// TIA Portal project "E95238_MCC1200_Sisecam_India" (V17)

(* hardware
DEVICE "S71500/ET200MP station_1"  S7-1500 station
   slot 0: "Rail_0"  Rack  6ES7 590-1***0-0AA0
   slot 1: "R150AP1"  CPU 1515-2 PN  6ES7 515-2AM02-0AB0  V2.8
      slot 3: "CPU display_1"  6ES7591-1BA00-0AA0
      slot 32768: "PROFINET_MCC1200"  X1
         slot 32769: "Port_1"  X1 P1
         slot 32770: "Port_2"  X1 P2
      slot 33024: "PCNETWORK_MCC1200"  X2
         slot 33025: "Port_1"  X2 P1
      slot 34817: "Virtual CP interface port_1"  Virtual CP interface port  Virtual CP interface port
   slot 2: "DI 16x24VDC HF_1"  DI 16x24VDC HF  6ES7 521-1BH00-0AB0  V2.2
DEVICE "ET 200SP station_2"  ET 200SP-Station
   slot 0: "Rack_0"  Rack  6ES5 710-8MAx1
   slot 0: "R195AP1"  IM 155-6 PN ST  6ES7 155-6AU01-0BN0  V4.1
   slot 1: "MasterCounter"  TM PosInput 1  6ES7 138-6BA00-0BA0  V1.3
      slot 1: "MasterCounter"  TM PosInput 1
   slot 2: "TM PosInput 1_2"  TM PosInput 1  6ES7 138-6BA00-0BA0  V1.3
      slot 1: "TM PosInput 1_2"  TM PosInput 1
   slot 3: "TM PosInput 1_3"  TM PosInput 1  6ES7 138-6BA00-0BA0  V1.2
      slot 1: "TM PosInput 1_3"  TM PosInput 1
   slot 4: "DI 16x24VDC ST_4"  DI 16x24VDC ST  6ES7 131-6BH01-0BA0  V0.0
      slot 1: "DI 16x24VDC ST_4"  DI 16x24VDC ST
   slot 5: "DI 16x24VDC ST_1"  DI 16x24VDC ST  6ES7 131-6BH01-0BA0  V0.0
      slot 1: "DI 16x24VDC ST_1"  DI 16x24VDC ST
   slot 6: "DI 16x24VDC ST_5"  DI 16x24VDC ST  6ES7 131-6BH01-0BA0  V0.0
      slot 1: "DI 16x24VDC ST_5"  DI 16x24VDC ST
   slot 7: "DQ 16x24VDC/0.5A ST_1"  DQ 16x24VDC/0.5A ST  6ES7 132-6BH01-0BA0  V0.0
      slot 1: "DQ 16x24VDC/0.5A ST_1"  DQ 16x24VDC/0.5A ST
   slot 8: "DQ 16x24VDC/0.5A ST_2"  DQ 16x24VDC/0.5A ST  6ES7 132-6BH01-0BA0  V0.0
      slot 1: "DQ 16x24VDC/0.5A ST_2"  DQ 16x24VDC/0.5A ST
   slot 9: "Server module_1"  Server module  6ES7 193-6PA00-0AA0  V1.1
      slot 1: "Server module_1"  Server module
   slot 127: "BA 2xRJ45"  BA 2xRJ45  6ES7 193-6AR00-0AA0  V0.0
      slot 1: "Port_1"  X1 P1 R  6ES7 193-6AR00-0AA0  V0.0
      slot 2: "Port_2"  X1 P2 R  6ES7 193-6AR00-0AA0  V0.0
DEVICE "ET 200SP station_1"  ET 200SP-Station
   slot 0: "Telaio di montaggio_0"  Rack  6ES5 710-8MAx1
   slot 1: "2B160AP"  CPU 1512SP-1 PN  6ES7 512-1DK01-0AB0  V2.9
      slot 32768: "PROFINET_YC2"  X1
   slot 2: "TM PosInput 1_1"  TM PosInput 1  6ES7 138-6BA00-0BA0  V1.2
      slot 1: "TM PosInput 1_1"  TM PosInput 1
   slot 3: "DI 16x24VDC ST_1"  DI 16x24VDC ST  6ES7 131-6BH01-0BA0  V0.0
      slot 1: "DI 16x24VDC ST_1"  DI 16x24VDC ST
   slot 4: "DI 8x24VDC ST_1"  DI 8x24VDC ST  6ES7 131-6BF01-0BA0  V0.0
      slot 1: "DI 8x24VDC ST_1"  DI 8x24VDC ST
   slot 5: "DQ 8x24VDC/0.5A ST_1"  DQ 8x24VDC/0.5A ST  6ES7 132-6BF01-0BA0  V0.0
      slot 1: "DQ 8x24VDC/0.5A ST_1"  DQ 8x24VDC/0.5A ST
   slot 6: "DQ 8x24VDC/0.5A ST_2"  DQ 8x24VDC/0.5A ST  6ES7 132-6BF01-0BA0  V0.0
      slot 1: "DQ 8x24VDC/0.5A ST_1"  DQ 8x24VDC/0.5A ST
   slot 7: "AQ 4xU/I ST_1"  AQ 4xU/I ST  6ES7 135-6HD00-0BA1  V1.1
      slot 1: "AQ 4xU/I ST_1"  AQ 4xU/I ST
   slot 8: "AQ 4xU/I ST_2"  AQ 4xU/I ST  6ES7 135-6HD00-0BA1  V1.1
      slot 1: "AQ 4xU/I ST_2"  AQ 4xU/I ST
   slot 9: "Modulo server_1"  Server module  6ES7 193-6PA00-0AA0  V1.1
      slot 1: "Modulo server_1"  Server module
   slot 127: "BA 2xRJ45"  BA 2xRJ45  6ES7 193-6AR00-0AA0  V0.0
      slot 32769: "Port_1"  6ES7 193-6AR00-0AA0
      slot 32770: "Port_2"  6ES7 193-6AR00-0AA0
DEVICE "GSD device_1"  GSD.Device.PN
   slot 0: "Rack"  Rack  V1.0
   slot 0: "Y2B412AP1"  55130 IMPACT67 DIO16 IRT  55130  1.02.00
      slot 0: "55130 IMPACT67 DIO16 IRT_1"  55130 IMPACT67 DIO16 IRT
      slot 1: "55130 IMPACT67 DIO16 IRT"  55130 IMPACT67 DIO16 IRT
         slot 1: "Port 1"  Port 1
         slot 2: "Port 2"  Port 2
      slot 1: "Device_1"  Device
         slot 0: "Parameter/Diagnostic"  Parameter/Diagnostic
         slot 1: "Digital IO"  Digital IO
DEVICE "GSD device_3"  GSD.Device.PN
   slot 0: "Rack"  Rack  V1.0
   slot 0: "Y2B411AP1"  55130 IMPACT67 DIO16 IRT  55130  1.02.00
      slot 0: "55130 IMPACT67 DIO16 IRT_1"  55130 IMPACT67 DIO16 IRT
      slot 1: "55130 IMPACT67 DIO16 IRT"  55130 IMPACT67 DIO16 IRT
         slot 1: "Port 1"  Port 1
         slot 2: "Port 2"  Port 2
      slot 1: "Device_1"  Device
         slot 0: "Parameter/Diagnostic"  Parameter/Diagnostic
         slot 1: "Digital IO"  Digital IO
DEVICE "GSD device_4"  GSD.Device.PN
   slot 0: "Rack"  Rack  V1.0
   slot 0: "Y2B413AP1"  55130 IMPACT67 DIO16 IRT  55130  1.02.00
      slot 0: "55130 IMPACT67 DIO16 IRT_1"  55130 IMPACT67 DIO16 IRT
      slot 1: "55130 IMPACT67 DIO16 IRT"  55130 IMPACT67 DIO16 IRT
         slot 1: "Port 1"  Port 1
         slot 2: "Port 2"  Port 2
      slot 1: "Device_1"  Device
         slot 0: "Parameter/Diagnostic"  Parameter/Diagnostic
         slot 1: "Digital IO"  Digital IO
DEVICE "GSD device_5"  GSD.Device.PN
   slot 0: "Rack"  Rack  V1.0
   slot 0: "Y2B414AP1"  55130 IMPACT67 DIO16 IRT  55130  1.02.00
      slot 0: "55130 IMPACT67 DIO16 IRT_1"  55130 IMPACT67 DIO16 IRT
      slot 1: "55130 IMPACT67 DIO16 IRT"  55130 IMPACT67 DIO16 IRT
         slot 1: "Port 1"  Port 1
         slot 2: "Port 2"  Port 2
      slot 1: "Device_1"  Device
         slot 0: "Parameter/Diagnostic"  Parameter/Diagnostic
         slot 1: "Digital IO"  Digital IO
DEVICE "GSD device_7"  GSD.Device.PN
   slot 0: "Rack"  Rack  V1.0
   slot 0: "Y2B415AP1"  55130 IMPACT67 DIO16 IRT  55130  1.02.00
      slot 0: "55130 IMPACT67 DIO16 IRT_1"  55130 IMPACT67 DIO16 IRT
      slot 1: "55130 IMPACT67 DIO16 IRT"  55130 IMPACT67 DIO16 IRT
         slot 1: "Port 1"  Port 1
         slot 2: "Port 2"  Port 2
      slot 1: "Device_1"  Device
         slot 0: "Parameter/Diagnostic"  Parameter/Diagnostic
         slot 1: "Digital IO"  Digital IO
DEVICE "ET 200SP station_3"  ET 200SP-Station
   slot 0: "Telaio di montaggio_0"  Rack  6ES5 710-8MAx1
   slot 1: "1B160AP"  CPU 1512SP-1 PN  6ES7 512-1DK01-0AB0  V2.9
      slot 32768: "PROFINET_YC1"  X1
   slot 2: "TM PosInput 1_1"  TM PosInput 1  6ES7 138-6BA00-0BA0  V1.2
      slot 1: "TM PosInput 1_1"  TM PosInput 1
   slot 3: "DI 16x24VDC ST_1"  DI 16x24VDC ST  6ES7 131-6BH01-0BA0  V0.0
      slot 1: "DI 16x24VDC ST_1"  DI 16x24VDC ST
   slot 4: "DI 8x24VDC ST_1"  DI 8x24VDC ST  6ES7 131-6BF01-0BA0  V0.0
      slot 1: "DI 8x24VDC ST_1"  DI 8x24VDC ST
   slot 5: "DI 16x24VDC ST_2"  DI 16x24VDC ST  6ES7 131-6BH01-0BA0  V0.0
      slot 1: "DI 16x24VDC ST_2"  DI 16x24VDC ST
   slot 6: "DQ 8x24VDC/0.5A ST_1"  DQ 8x24VDC/0.5A ST  6ES7 132-6BF01-0BA0  V0.0
      slot 1: "DQ 8x24VDC/0.5A ST_1"  DQ 8x24VDC/0.5A ST
   slot 7: "DQ 16x24VDC/0.5A ST_1"  DQ 16x24VDC/0.5A ST  6ES7 132-6BH01-0BA0  V0.0
      slot 1: "DQ 16x24VDC/0.5A ST_1"  DQ 16x24VDC/0.5A ST
   slot 8: "AQ 4xU/I ST_1"  AQ 4xU/I ST  6ES7 135-6HD00-0BA1  V1.1
      slot 1: "AQ 4xU/I ST_1"  AQ 4xU/I ST
   slot 9: "AQ 4xU/I ST_2"  AQ 4xU/I ST  6ES7 135-6HD00-0BA1  V1.1
      slot 1: "AQ 4xU/I ST_2"  AQ 4xU/I ST
   slot 10: "Modulo server_1"  Server module  6ES7 193-6PA00-0AA0  V1.1
      slot 1: "Modulo server_1"  Server module
   slot 127: "BA 2xRJ45"  BA 2xRJ45  6ES7 193-6AR00-0AA0  V0.0
      slot 32769: "Port_1"  6ES7 193-6AR00-0AA0
      slot 32770: "Port_2"  6ES7 193-6AR00-0AA0
DEVICE "GSD device_9"  GSD.Device.PN
   slot 0: "Rack"  Rack  V1.0
   slot 0: "Y1B415AP1"  55130 IMPACT67 DIO16 IRT  55130  1.02.00
      slot 0: "55130 IMPACT67 DIO16 IRT_1"  55130 IMPACT67 DIO16 IRT
      slot 1: "55130 IMPACT67 DIO16 IRT"  55130 IMPACT67 DIO16 IRT
         slot 1: "Port 1"  Port 1
         slot 2: "Port 2"  Port 2
      slot 1: "Device_1"  Device
         slot 0: "Parameter/Diagnostic"  Parameter/Diagnostic
         slot 1: "Digital IO"  Digital IO
DEVICE "GSD device_10"  GSD.Device.PN
   slot 0: "Rack"  Rack  V1.0
   slot 0: "Y1B414AP1"  55130 IMPACT67 DIO16 IRT  55130  1.02.00
      slot 0: "55130 IMPACT67 DIO16 IRT_1"  55130 IMPACT67 DIO16 IRT
      slot 1: "55130 IMPACT67 DIO16 IRT"  55130 IMPACT67 DIO16 IRT
         slot 1: "Port 1"  Port 1
         slot 2: "Port 2"  Port 2
      slot 1: "Device_1"  Device
         slot 0: "Parameter/Diagnostic"  Parameter/Diagnostic
         slot 1: "Digital IO"  Digital IO
DEVICE "GSD device_11"  GSD.Device.PN
   slot 0: "Rack"  Rack  V1.0
   slot 0: "Y1B413AP1"  55130 IMPACT67 DIO16 IRT  55130  1.02.00
      slot 0: "55130 IMPACT67 DIO16 IRT_1"  55130 IMPACT67 DIO16 IRT
      slot 1: "55130 IMPACT67 DIO16 IRT"  55130 IMPACT67 DIO16 IRT
         slot 1: "Port 1"  Port 1
         slot 2: "Port 2"  Port 2
      slot 1: "Device_1"  Device
         slot 0: "Parameter/Diagnostic"  Parameter/Diagnostic
         slot 1: "Digital IO"  Digital IO
DEVICE "GSD device_13"  GSD.Device.PN
   slot 0: "Rack"  Rack  V1.0
   slot 0: "Y1B412AP1"  55130 IMPACT67 DIO16 IRT  55130  1.02.00
      slot 0: "55130 IMPACT67 DIO16 IRT_1"  55130 IMPACT67 DIO16 IRT
      slot 1: "55130 IMPACT67 DIO16 IRT"  55130 IMPACT67 DIO16 IRT
         slot 1: "Port 1"  Port 1
         slot 2: "Port 2"  Port 2
      slot 1: "Device_1"  Device
         slot 0: "Parameter/Diagnostic"  Parameter/Diagnostic
         slot 1: "Digital IO"  Digital IO
DEVICE "GSD device_14"  GSD.Device.PN
   slot 0: "Rack"  Rack  V1.0
   slot 0: "Y1B411AP1"  55130 IMPACT67 DIO16 IRT  55130  1.02.00
      slot 0: "55130 IMPACT67 DIO16 IRT_1"  55130 IMPACT67 DIO16 IRT
      slot 1: "55130 IMPACT67 DIO16 IRT"  55130 IMPACT67 DIO16 IRT
         slot 1: "Port 1"  Port 1
         slot 2: "Port 2"  Port 2
      slot 1: "Device_1"  Device
         slot 0: "Parameter/Diagnostic"  Parameter/Diagnostic
         slot 1: "Digital IO"  Digital IO
DEVICE "GSD device_15"  GSD.Device.PN
   slot 0: "Rack"  Rack  V1.0
   slot 0: "Y1B416AP1"  55130 IMPACT67 DIO16 IRT  55130  1.02.00
      slot 0: "55130 IMPACT67 DIO16 IRT_1"  55130 IMPACT67 DIO16 IRT
      slot 1: "55130 IMPACT67 DIO16 IRT"  55130 IMPACT67 DIO16 IRT
         slot 1: "Port 1"  Port 1
         slot 2: "Port 2"  Port 2
      slot 1: "Device_1"  Device
         slot 0: "Parameter/Diagnostic"  Parameter/Diagnostic
         slot 1: "Digital IO"  Digital IO
DEVICE "GSD device_2"  GSD.Device.PN
   slot 0: "Rack"  Rack  V1.0
   slot 0: "Y1B417AP1"  55130 IMPACT67 DIO16 IRT  55130  1.02.00
      slot 0: "55130 IMPACT67 DIO16 IRT_1"  55130 IMPACT67 DIO16 IRT
      slot 1: "55130 IMPACT67 DIO16 IRT"  55130 IMPACT67 DIO16 IRT
         slot 1: "Port 1"  Port 1
         slot 2: "Port 2"  Port 2
      slot 1: "Device_1"  Device
         slot 0: "Parameter/Diagnostic"  Parameter/Diagnostic
         slot 1: "Digital IO"  Digital IO
DEVICE "GSD device_6"  GSD.Device.PN
   slot 0: "Rack"  Rack  V1.0
   slot 0: "Y1B418AP1"  55130 IMPACT67 DIO16 IRT  55130  1.02.00
      slot 0: "55130 IMPACT67 DIO16 IRT_1"  55130 IMPACT67 DIO16 IRT
      slot 1: "55130 IMPACT67 DIO16 IRT"  55130 IMPACT67 DIO16 IRT
         slot 1: "Port 1"  Port 1
         slot 2: "Port 2"  Port 2
      slot 1: "Device_1"  Device
         slot 0: "Parameter/Diagnostic"  Parameter/Diagnostic
         slot 1: "Digital IO"  Digital IO
DEVICE "GSD device_8"  GSD.Device.PN
   slot 0: "Rack"  Rack  V1.0
   slot 0: "Y2B418AP1"  55130 IMPACT67 DIO16 IRT  55130  1.02.00
      slot 0: "55130 IMPACT67 DIO16 IRT_1"  55130 IMPACT67 DIO16 IRT
      slot 1: "55130 IMPACT67 DIO16 IRT"  55130 IMPACT67 DIO16 IRT
         slot 1: "Port 1"  Port 1
         slot 2: "Port 2"  Port 2
      slot 1: "Device_1"  Device
         slot 0: "Parameter/Diagnostic"  Parameter/Diagnostic
         slot 1: "Digital IO"  Digital IO
DEVICE "GSD device_12"  GSD.Device.PN
   slot 0: "Rack"  Rack  V1.0
   slot 0: "Y2B417AP1"  55130 IMPACT67 DIO16 IRT  55130  1.02.00
      slot 0: "55130 IMPACT67 DIO16 IRT_1"  55130 IMPACT67 DIO16 IRT
      slot 1: "55130 IMPACT67 DIO16 IRT"  55130 IMPACT67 DIO16 IRT
         slot 1: "Port 1"  Port 1
         slot 2: "Port 2"  Port 2
      slot 1: "Device_1"  Device
         slot 0: "Parameter/Diagnostic"  Parameter/Diagnostic
         slot 1: "Digital IO"  Digital IO
DEVICE "GSD device_16"  GSD.Device.PN
   slot 0: "Rack"  Rack  V1.0
   slot 0: "Y2B416AP1"  55130 IMPACT67 DIO16 IRT  55130  1.02.00
      slot 0: "55130 IMPACT67 DIO16 IRT_1"  55130 IMPACT67 DIO16 IRT
      slot 1: "55130 IMPACT67 DIO16 IRT"  55130 IMPACT67 DIO16 IRT
         slot 1: "Port 1"  Port 1
         slot 2: "Port 2"  Port 2
      slot 1: "Device_1"  Device
         slot 0: "Parameter/Diagnostic"  Parameter/Diagnostic
         slot 1: "Digital IO"  Digital IO
DEVICE "GSD device_17"  GSD.Device.PN
   slot 0: "Telaio di montaggio"  Rack  V1.0
   slot 1: "d405ap1"  D405AP1  6ES7 512-1DK01-0AB0  V2.9
      slot 0: "InputCPU0"  InputCPU0
      slot 1: "OutputCPU0"  OutputCPU0
      slot 2: "Interface"  Interface
         slot 1: "Port 1"  Port 1
         slot 2: "Port 2"  Port 2
         slot 3: "Port 3"  Port 3
*)

// ===== PLC "R150AP1"  CPU 1515-2 PN =====

VAR_GLOBAL   // PLC tag table "Default tag table"
   "FirstScan" AT %M0.0 : Bool;
   "AlwaysTRUE" AT %M0.2 : Bool;
   "AlwaysFALSE" AT %M0.3 : Bool;
   "AlwaysOFF_Debug" AT %M10.0 : Bool;
   "o.R195AP1.R251KA1.EncoderCommutation" AT %Q120.0 : Bool;
   "i.R195AP1.R11QF2/3.PowerFailure230VAuxiliary" AT %I120.1 : Bool;
   "i.R195AP1.R18QF3.PowerFailure24V_Commands" AT %I120.6 : Bool;
   "i.R195AP1.R18QF4.PowerFailure24V_Input" AT %I120.7 : Bool;
   "i.R195AP1.R18AP1.Redundacy24VOk" AT %I120.5 : Bool;
   "i.R195AP1.M216B1.GlassPresenceOnEncoder#1M216" AT %I122.0 : Bool;
   "i.R195AP1.M216B2.GlassPresenceOnEncoder#2M216" AT %I122.1 : Bool;
   "i.R195AP1.R427SL1.MinimumLevelOilTank" AT %I122.3 : Bool;
   "i.R195AP1.R427SL2.MaximumLevelOilTank" AT %I122.4 : Bool;
   "i.R195AP1.M212SB4.DefectButtonClass3" AT %I123.3 : Bool;
   "i.R195AP1.M212SB3.QualityB1" AT %I123.2 : Bool;
   "i.R195AP1.M212SB5.DefectButtonClass4" AT %I123.4 : Bool;
   "i.R195AP1.SCANNER.ScannerOn" AT %I124.0 : Bool;
   "i.R195AP1.SCANNER.Scanner(1)" AT %I124.1 : Bool;
   "o.R195AP1.R251KA2.Jog" AT %Q120.1 : Bool;
   "o.R195AP1.R252HL1.SafetiesON" AT %Q121.1 : Bool;
   "o.R195AP1.R252HL2.EnableCPUA" AT %Q121.2 : Bool;
   "o.R195AP1.R252HL2.EnableCPUB" AT %Q121.3 : Bool;
   "o.R195AP1.R252KA1.SCANNER.RiseBreakingBar" AT %Q121.5 : Bool;
   "o.R195AP1.R252KA2.SCANNER.GlassToSQC" AT %Q121.6 : Bool;
   "o.R195AP1.M216YV1.DigitizerRise/descentEncoder1" AT %Q122.0 : Bool;
   "o.R195AP1.M216YV2.DigitizeRise/descentEncoder2" AT %Q122.1 : Bool;
   "o.R195AP1.R429YV1.StartFillingPumpCuttingTank" AT %Q122.5 : Bool;
   "o.R195AP1.M221YV2.UpperHolderControl" AT %Q122.7 : Bool;
   "o.R195AP1.M221YV1.BreakoutBarControl" AT %Q122.6 : Bool;
   "o.R195AP1.M221HL1.CutTrasversalBridge1" AT %Q123.1 : Bool;
   "o.R195AP1.M221HL2.CutTrasversalBridge2" AT %Q123.2 : Bool;
   "i.R195AP1.R125KA1CPU_A_Enabled" AT %I121.3 : Bool;
   "i.R195AP1.R125SA1SelectionOnCPU_B" AT %I121.4 : Bool;
   "i.R150AP1.Recognition CPU A" AT %I20.2 : Bool;
   "cigliutti" AT %M100.1 : Bool;
   "i.R195AP1.R18QF7.PowerSupply24VLogic" AT %I121.1 : Bool;
   "i.R195AP1.R427SSP1.CompressedAirPresenceCuttingBridge" AT %I122.5 : Bool;
   "i.R195AP1.R18QF8.PowerSupply24VLogic" AT %I121.2 : Bool;
   "i.R195AP1.M212SB1.DefectButtonClass3" AT %I123.0 : Bool;
   "i.R195AP1.M212SB2.DefectButtonClass4" AT %I123.1 : Bool;
   "o.R195AP1.A255KA6.Anomaly" AT %Q4.5 : Bool;
   "o.R195AP1.A257KA4.AllowM225" AT %Q6.3 : Bool;
   "o.R195AP1.A257KA5.AllowM225(1)" AT %Q6.4 : Bool;
   "o.R195AP1.A252KA3.SCANNER.NoGlassBreak" AT %Q121.7 : Bool;
   "o.R195AP1.M212SB3.M212SB6.GlassRequestQlt" AT %Q123.0 : Bool;
   "o.R195AP1.FanRotationM250" AT %Q2.0 : Bool;
   "i.MCC1256B1_IDevice" AT %I2500.0 : "UDT_YCut_IdeviceFromBridge";
   "i_HSCInput_Count1" AT %I30.0 : "LPD_typeCountFeedbackCh";
   "i_HSCInput_Count2" AT %I160.0 : "LPD_typeCountFeedbackCh";
   "i_HSCInput_Count3" AT %I180.0 : "LPD_typeCountFeedbackCh";
   "i.MCC1256B2_IDevice" AT %I3000.0 : "UDT_YCut_IdeviceFromBridge";
   "i_IDeviceFromZ300" AT %I3300.0 : "UDT_iDeviceZ301--->Z200";
   "o_HSCOutput_Count1" AT %Q30.0 : "LPD_typeCountControlCh";
   "o_HSCOutput_Count2" AT %Q160.0 : "LPD_typeCountControlCh";
   "o_HSCOutput_Count3" AT %Q180.0 : "LPD_typeCountControlCh";
   "o.MCC1256B1_IDevice" AT %Q2500.0 : "UDT_YCut_IdeviceToBridge";
   "o.MCC1256B2_IDevice" AT %Q3000.0 : "UDT_YCut_IdeviceToBridge";
   "o_IDeviceToZ300_INO" AT %Q3300.0 : "UDT_iDeviceZ301<---Z200_INO";
   "TestTag64" AT %M2.0 : LInt;
   "i.R195AP1.R18QF1.PowerFailure24VSuplly1" AT %I120.3 : Bool;
   "i.R195AP1.R18QF2.PowerFailure24VSuplly2" AT %I120.4 : Bool;
   "i.R150AP1.Selected CPU B" AT %I20.1 : Bool;
   "i.R150AP1.Selected CPU A" AT %I20.0 : Bool;
   "i.R150AP1.Anomay Power supply  CPU B" AT %I20.3 : Bool;
   "salto" AT %MW12 : Int;
   "Berg_Check" AT %M775.0 : Bool;
   "o.R195AP1.M221HL3.CutTrasversalBridge3" AT %Q123.3 : Bool;
   "o.R195AP1.R254KA1.BrandingMachineAllow" AT %Q123.5 : Bool;
   "o.R195AP1.R254KA2.BrandingMachineAllow" AT %Q123.6 : Bool;
   "o.R195AP1.R254KA3.BrandingMachineAllow" AT %Q123.7 : Bool;
   "i.R195AP1.SCANNER.Scanner(2)" AT %I124.2 : Bool;
   "i.R195AP1.SCANNER.Scanner(3)" AT %I124.3 : Bool;
   "o.R195AP1.R251KA3.CpuASerSel" AT %Q120.3 : Bool;
   "o.R195AP1.R251KA4.CpuBSerSel" AT %Q120.4 : Bool;
   "o.R195AP1.R251KA5.IsraRiseBreakBar" AT %Q120.5 : Bool;
   "o.R195AP1.R251KA6.IsraSheetToQlt" AT %Q120.6 : Bool;
   "prova" AT %I3576.0 : Bool;
   "i.MCC1204_IDeviceFromMarkers" AT %I3500.0 : "UDT_Marker_IDeviceFromBridge";
   "o.MCC1204_IDeviceToMarkers" AT %Q3500.0 : "UDT_Marker_IDeviceToBridge";
   "Check" AT %M1.0 : Bool;
   "o_IDeviceToZ300OUT" AT %A3304.0 : "UDT_iDevice_MCC1201<---Mcc1200_OUT";
END_VAR

VAR_GLOBAL CONSTANT   // PLC tag table "Default tag table"
   "DSTRSIZEDESCR" : DInt := 30;   // Default size of the description string
   "DMAXYCUTBRIDGE" : DInt := 2;   // Number of YCUT bridges
   "DMAXYCUTBRIDGE_IND" : DInt := 1;   // Number of YCUT bridges -1 used for index
   "DMAXYHEADS" : DInt := 16;   // Number of YCUT heads
   "DMAXYHEADS_IND" : DInt := 15;   // Number of YCUT heads -1 used for index
   "DMAXXHEADS" : DInt := 5;   // Number of XCUT bridge
   "DMAXXHEADS_IND" : DInt := 4;   // Number of XCUT bridge -1 used for index
   "DMAXLITE" : DInt := 12;   // Number of lites
   "DMAXLITE_IND" : DInt := 11;   // Number of lites -1 used for index
   "DMAXSEPROLLBANK" : DInt := 4;   // Number of separotor roll bank
   "DMAXSEPROLLBANK_IND" : DInt := 3;   // Number of separator roll bank -1 used for index
   "DMAXPROTLAYER" : DInt := 8;   // Number of protection layer
   "DMAXPROTLAYER_IND" : DInt := 7;   // Number of protection layer -1 used for index
   "DSTRSIZEDEFID" : DInt := 50;   // Default size of the defect ID size
   "DNUMDEFEXT" : DInt := 10000;   // Maximum number of defect extended on buffer
   "DNUMDEFEXT_IND" : DInt := 9999;   // Maximum number of defect extended on buffer -1 used for index
   "DMAXNUMCLASS" : DInt := 30;   // Maximum number of defect classes
   "DMAXNUMCLASS_IND" : DInt := 29;   // Maximum number of defect classes -1 used for index
   "DMAXNUMDEFCLASS" : DInt := 500;   // Maximum number of defect for classes
   "DMAXNUMDEFCLASS_IND" : DInt := 499;   // Maximum number of defect for classes -1 used for index
   "DMAXDEFECTID" : DInt := 2000000000;   // Maximum ID defect
   "DMAXTRACKCAP" : DInt := 50;   // Maximum number of caps on tracking
   "DMAXTRACKCAP_IND" : DInt := 49;   // Maximum number of caps on tracking -1 used for index
   "DMAXTRACKMACHINE" : DInt := 32;   // Maximum number of machine on tracking
   "DMAXTRACKMACHINE_IND" : DInt := 31;   // Maximum number of machine on tracking -1 used for index
   "DMAXPLATEID" : DInt := 2000000000;   // Maximum ID plate
   "DMAXELEMWAKEUPNEWPLATE" : DInt := 16;   // Maximum number of element to wakeup new plate
   "DMAXELEMWAKEUPNEWPLATE_IND" : DInt := 15;   // Maximum number of element to wakeup new plate -1 used for index
   "DMACHINEINDEX_LASTOPTLINE" : DInt := 0;   // Position index on the machine tracking of the last optimization line
   "DMACHINEINDEX_YCUT1" : DInt := 1;   // Position index on the machine tracking of the last YCUT#1
   "DMACHINEINDEX_YCUT2" : DInt := 2;   // Position index on the machine tracking of the last YCUT#2
   "DMACHINEINDEX_XCUT1" : DInt := 3;   // Position index on the machine tracking of the last XCUT#1
   "DMACHINEINDEX_XCUT2" : DInt := 4;   // Position index on the machine tracking of the last XCUT#2
   "DMACHINEINDEX_XCUT3" : DInt := 5;   // Position index on the machine tracking of the last XCUT#3
   "DMACHINEINDEX_XCUT4" : DInt := 6;   // Position index on the machine tracking of the last XCUT#4
   "DMACHINEINDEX_XCUT5" : DInt := 7;   // Position index on the machine tracking of the last XCUT#5
   "DMACHINEINDEX_SNAPROLL" : DInt := 8;   // Position index on the machine tracking of the snaproll
   "DMINLEHRSPEED_MM_MIN" : DInt := 500;   // Minimum lehr speed [mm/min]
   "DMAXLEHRSPEED_MM_MIN" : DInt := 25000;   // Maximum lehr speed [mm/min]
   "DCULLETDESTMASK" : LInt := 1099511627776;   // Cullet destination mask [mask]
   "DQUALITYDESTMASK1" : LInt := 512;   // Quality 1 destination mask [mask]
   "DMAXELEMTRACKSEARCH" : DInt := 20;   // Maximum number of element on tracking search
   "DMAXELEMTRACKSEARCH_IND" : DInt := 19;   // Maximum number of element on tracking search -1 used for index
   "CONNUOC_DIGITIZER_1" : Conn_Ouc := 16#1;   // Connection ID for serial converter FM152-1
   "IPV4_DIGITIZER_1_IP1" : Byte := 192;   // IP_1 for serial converter FM152-1
   "IPV4_DIGITIZER_1_IP2" : Byte := 168;   // IP_2 for serial converter FM152-1
   "IPV4_DIGITIZER_1_IP3" : Byte := 20;   // IP_3 for serial converter FM152-1
   "IPV4_DIGITIZER_1_IP4" : Byte := 12;   // IP_4 for serial converter FM152-1
   "UINT_DIGIITZER_1_PORT" : UInt := 4001;   // Port for serial converter Fm152-1
   "CONNUOC_DIGITIZER_2" : Conn_Ouc := 16#2;   // Connection ID for serial converter FM152-2
   "IPV4_DIGITIZER_2_IP1" : Byte := 192;   // IP_1 for serial converter FM152-2
   "IPV4_DIGITIZER_2_IP2" : Byte := 168;   // IP_2 for serial converter FM152-2
   "IPV4_DIGITIZER_2_IP3" : Byte := 20;   // IP_3 for serial converter FM152-2
   "IPV4_DIGITIZER_2_IP4" : Byte := 13;   // IP_4 for serial converter FM152-2
   "UINT_DIGIITZER_2_PORT" : UInt := 4001;   // Port for serial converter Fm152-2
   "DINDEXNEWCAPAVAILABLE_YCUT1" : UInt := 0;   // Index for new cap available for YCUT1
   "DINDEXNEWCAPAVAILABLE_YCUT2" : UInt := 1;   // Index for new cap available for YCUT2
   "CONNANY_YCUT1_ID" : Conn_Any := 16#100;   // Connection ID for YCUT#1
   "CONNANY_YCUT2_ID" : Conn_Any := 16#101;   // Connection ID for YCUT#2
   "DMAXMARKERMISSIONONTANK" : DInt := 99;   // Maximum number of mission on marker tank
   "DMAXMARKERMISSIONSEND" : DInt := 19;   // Maximum number of mission to send to marker tank
   "DNUMBEROFDESTINATION_Z300" : DInt := 63;   // Number of destination -1
   "DMAXLENGHTCONVOY_CMM" : DInt := 630000;   // Maximum lenght convoy [mm/100]
   "DMAXCAP_Z300" : DInt := 2;   // Maximum number of caps Z300
   "DMACHINEINDEX_Z300" : DInt := 9;   // Position index on the machine tracking of the Z300
   "CONNANY_MARKER_ID" : Conn_Any := 16#102;   // Connection ID for Marker
   "CONNANY_Z300_ID" : Conn_Any := 16#103;   // Connection ID for Z300
   "CONNUOC_BPS_SERVERA" : Conn_Ouc := 16#3;   // Connection ID for BPS Server A
   "IPV4_BPS_SERVERA_IP1" : Byte := 192;   // IP_1 for BPS Server A
   "IPV4_BPS_SERVERA_IP2" : Byte := 168;   // IP_2 for BPS Server A
   "IPV4_BPS_SERVERA_IP3" : Byte := 100;   // IP_3 for BPS Server A
   "IPV4_BPS_SERVERA_IP4" : Byte := 3;   // IP_4 for BPS Server A
   "UINT_BPS_SERVERA_PORT" : UInt := 6000;   // Port for BPS Server A
   "SIMULATION_ACTIVE" : Bool := 1;   // Enable simulation
   "DNUMDEFFOROPT" : DInt := 11;   // Maximum number of defect for optimizer
   "DNUMDEFFOROPT_IND" : DInt := 10;   // Maximum number of defect for optimizer -1 used for index
   "DNUMDEFFORREPORT" : DInt := 10;   // Maximum number of defect for report
   "DNUMDEFFORREPORT_IND" : DInt := 9;   // Maximum number of defect for report -1 used for index
   "CONNUOC_OPTIMIZER_SMALLPCK" : Conn_Ouc := 16#5;   // Connection ID for optimizer small packet port
   "CONNUOC_OPTIMIZER_BIGPCK" : Conn_Ouc := 16#6;   // Connection ID for optimizer big packet port
   "UINT_OPTIMIZER_PORT_SMALLPCK" : UInt := 7000;   // Port for optimizer small packet
   "UINT_OPTIMIZER_PORT_BIGPCK" : UInt := 7001;   // Port for optimizer big packet
   "DMAXNUMMESSAGETANK" : DInt := 200;   // Number of messages on tank
   "DMAXNUMMESSAGETANK_IND" : DInt := 199;   // Number of messages on tank index (Always -1)
   "DCULLETCAUSE_XCUTMISSING" : DInt := 200;   // Cullet cause - X Cut missing
   "DCULLETCAUSE_YCUTMISSING" : DInt := 201;   // Cullet cause - Y Cut missing generic
   "DCULLETCAUSE_MARKMISSING" : DInt := 202;   // Cullet cause - Mark missing
   "DCULLETCAUSE_BPMREDEST" : DInt := 203;   // Cullet cause - BPM Operator redestination
   "DCULLETCAUSE_YCUTMISSING_GLASSBREAK" : DInt := 204;   // Cullet cause - Glass break
   "DCULLETCAUSE_YCUTMISSING_OPERHEADDIS" : DInt := 205;   // Cullet cause - Operator head disabled
   "DCULLETCAUSE_YCUTMISSING_BRIDGEANOMALY" : DInt := 206;   // Cullet cause - Bridge anomaly
   "DCULLETCAUSE_Z200_CLEAN" : DInt := 207;   // Cullet cause - Z200 cleaning
   "DCULLETCAUSE_THICK_OUTRANGE" : DInt := 208;   // Cullet cause - Thickness outside range
   "DCULLETCAUSE_CAPDATATIMEOUT" : DInt := 209;   // Cullet cause - Cap data timeout
   "DEVENTS_REDESTINATION" : DInt := 30;   // Events - Redestination message
   "DEVENTS_CULLETDESTINATION" : DInt := 200;   // Events - Cullet destination
   "DEVENTS_MARKER_MISSION" : DInt := 80;   // Events - Markers mission
   "DMAXGLASSBREAKMACHINE" : DInt := 5;   // Maximum number of glass break machine
   "DMAXGLASSBREAKMACHINE_IND" : DInt := 4;   // Maximum number of glass break machine index (Always -1)
   "DMAXGLASSBREAKSECTORS" : DInt := 300;   // Maximum number of glass break sectors
   "DMAXGLASSBREAKSECTORS_IND" : DInt := 299;   // Maximum number of glass break sectors index (Always -1)
   "DMAXGLASSDATASECTORS" : DInt := 300;   // Maximum number of glass data sectors
   "DMAXGLASSDATASECTORS_IND" : DInt := 299;   // Maximum number of glass data sectors index (Always -1)
   "DMAXGLASSDATAMACHINE" : DInt := 5;   // Maximum number of glass data machine
   "DMAXGLASSDATAMACHINE_IND" : DInt := 4;   // Maximum number of glass data machine index (Always -1)
   "DEVENTS_REDEST_OPT" : DInt := 60;   // Events - Redestination from OPT
   "DMAXGLASSBREAKPHOTOCELL" : DInt := 32;   // Maximum number of glass break photocell
   "DMAXGLASSBREAKPHOTOCELL_IND" : DInt := 31;   // Maximum number of glass break photocell index (Always -1)
   "DMAXGLASSBREAKREQUEST" : DInt := 16;   // Maximum number of glass break request
   "DMAXGLASSBREAKREQUEST_IND" : DInt := 15;   // Maximum number of glass break request index (Always -1)
   "DMAXGLASSDATAREQUEST" : DInt := 16;   // Maximum number of glass data request
   "DMAXGLASSDATAREQUEST_IND" : DInt := 15;   // Maximum number of glass data request index (Always -1)
   "DMAXMARKERS" : DInt := 4;   // Maximum number of markers
   "DMAXMARKERS_IND" : DInt := 3;   // Maximum number of markers index (Always -1)
   "DGLASSBREAKMACHINEINDEX_M202" : DInt := 0;   // Glass break machine M202_Photocell_bridge
   "DGLASSBREAKMACHINEINDEX_M216" : DInt := 1;   // Glass break machine M216_digitizer
   "DGLASSBREAKMACHINEINDEX_M204" : DInt := 2;   // Glass break machine M204_drop_conv
   "DGLASSDATAMACHINEINDEX_MANUAL" : DInt := 0;   // Glass data machine MANUAL
   "DGLASSDATAMACHINEINDEX_SCANNER" : DInt := 1;   // Glass data machine SCANNER
   "DGLASSDATAMACHINEINDEX_CAMERA" : DInt := 2;   // Glass data machine CAMERA
   "DGLASSDATAGET_OPTMANAGERFB" : DInt := 0;   // Glass data get index
   "DGLASSDATAUPD_OPTMANAGERFB" : DInt := 0;   // Glass data update index (Manual machine)
   "DGLASSDATAUPD_ISRA5DFB" : DInt := 1;   // Glass data update index (Scanner machine)
   "CONNUOC_ISRA5D" : Conn_Ouc := 16#7;   // Connection ID for ISRA 5D
   "UINT_ISRA5D_PORT" : UInt := 4000;   // Port for ISRA5D
   "DGLASSBREAKGET_ISRA5DFB" : DInt := 10;   // Glass break get index (ISRA 5D)
   "COLDBACKUP_CONNUOC_SEND" : Conn_Ouc := 16#8;   // Connection ID for Cold Backup send
   "COLDBACKUP_CONNUOC_RECV" : Conn_Ouc := 16#9;   // Connection ID for Cold backup receive
   "COLDBACKUP_REMOTE_PORTSEND" : DInt := 7500;   // Port for cold backup send
   "COLDBACKUP_REMOTE_PORTRECV" : DInt := 7500;   // Port for cold backup receive
   "IPV4_BPS_SERVERB_IP1" : Byte := 192;   // IP_1 for BPS Server B
   "IPV4_BPS_SERVERB_IP2" : Byte := 168;   // IP_2 for BPS Server B
   "IPV4_BPS_SERVERB_IP3" : Byte := 100;   // IP_3 for BPS Server B
   "IPV4_BPS_SERVERB_IP4" : Byte := 4;   // IP_4 for BPS Server B
   "UINT_BPS_SERVERB_PORT" : UInt := 6000;   // Port for BPS Server B
   "CONNUOC_BPS_SERVERB" : Conn_Ouc := 16#4;   // Connection ID for BPS Server B
   "DGLASSBREAKGET_YCUT1" : DInt := 0;   // Glass break get index (YCUT 1)
   "DGLASSBREAKGET_YCUT2" : DInt := 1;   // Glass break get index (YCUT 2)
   "DGLASSBREAKGET_XCUT1" : DInt := 3;   // Glass break get index (XCUT 1)
   "DGLASSBREAKGET_XCUT2" : DInt := 4;   // Glass break get index (XCUT 2)
   "DGLASSBREAKGET_XCUT3" : DInt := 5;   // Glass break get index (XCUT 3)
   "DGLASSBREAKGET_XCUT4" : DInt := 6;   // Glass break get index (XCUT 4)
   "DGLASSBREAKGET_MARKER" : DInt := 7;   // Glass break get index (XCUT 5)
   "DQUALITYDESTMASK2" : LInt := 1048576;   // Quality 2 destination mask [mask]
   "DQUALITYDESTMASK3" : LInt := 2147483648;   // Quality 3 destination mask [mask]
   "CONNUOC_XCUT1" : Conn_Ouc := 16#10;   // Connection ID for modbus Xcut #1
   "IPV4_THICKNESS_IP1" : Byte := 192;   // IP_1 for serial converter thickness
   "IPV4_THICKNESS_IP2" : Byte := 168;   // IP_2 for serial converter thickness
   "IPV4_THICKNESS_IP3" : Byte := 21;   // IP_3 for serial converter thickness
   "IPV4_THICKNESS_IP4" : Byte := 202;   // IP_4 for serial converter thickness
   "UINT_THICKNESS_PORT" : UInt := 4000;   // Port for serial converter thickness
   "DMACHINEINDEX_ISRASNAP" : DInt := 10;   // Position index on the machine tracking of the isra signal
   "DEVENTS_TRAPSTATUS" : DInt := 44;   // Events - Trap status
   "DSTATUS_TRAPUP" : DInt := 21;   // Status - Trap UP
   "DSTATUS_TRAPDW" : DInt := 20;   // Status - Trap DW
   "DSTATUS_TRAP_AVAILABLE" : DInt := 3;   // Status - Trap available
   "DSTATUS_TRAP_OUTSERVICE" : DInt := 1;   // Status - Trap out of service
   "DMACHINE_TRAP_T1" : DInt := 201;   // Machine - Trap T1 Identifier
   "DEVENTS_CULLETLENGTH" : DInt := 45;   // Events - Cullet length
   "DCULLETTYPE_STRIPE" : DInt := 1;   // Cullet Type - Stripe
   "DMACHINE_TRAP_STRIPE" : DInt := 202;   // Machine - Trap stripe
   "DEVENTS_DESTSTATUS" : DInt := 41;
   "DEVENTS_DESTSTATUS_OUTSERVICE" : DInt := 1;
   "DEVENTS_DESTSTATUS_NOTAVAIL" : DInt := 2;
   "DEVENTS_DESTSTATUS_AVAILABLE" : DInt := 3;
   "DEVENTS_PLATE_STACKED" : DInt := 1;
   "DEVENTS_PLATE_REENTRY" : DInt := 2;
   "DEVENTS_PLATE_BROKEN" : DInt := 3;
   "DEVENTS_RACK_START" : DInt := 10;
   "DEVENTS_PACK_START" : DInt := 11;
   "DEVENTS_RACK_END" : DInt := 12;
   "DEVENTS_PACK_END" : DInt := 13;
   "DEVENTS_DEST_STATUS" : DInt := 41;
   "IPV4_XCUT1_IP1" : Byte := 192;   // IP_1 for Xcut #1
   "IPV4_XCUT1_IP2" : Byte := 168;   // IP_2 for Xcut #1
   "IPV4_XCUT1_IP3" : Byte := 20;   // IP_3 for Xcut #1
   "IPV4_XCUT1_IP4" : Byte := 111;   // IP_4 for Xcut #1
   "IPV4_XCUT2_IP1" : Byte := 192;   // IP_1 for Xcut #2
   "IPV4_XCUT2_IP2" : Byte := 168;   // IP_2 for Xcut #2
   "IPV4_XCUT2_IP3" : Byte := 20;   // IP_3 for Xcut #2
   "IPV4_XCUT2_IP4" : Byte := 112;   // IP_4 for Xcut #2
   "IPV4_XCUT3_IP1" : Byte := 192;   // IP_1 for Xcut #3
   "IPV4_XCUT3_IP2" : Byte := 168;   // IP_2 for Xcut #3
   "IPV4_XCUT3_IP3" : Byte := 20;   // IP_3 for Xcut #3
   "IPV4_XCUT3_IP4" : Byte := 113;   // IP_4 for Xcut #3
   "CONNUOC_XCUT2" : Conn_Ouc := 16#11;   // Connection ID for modbus Xcut #2
   "CONNUOC_XCUT3" : Conn_Ouc := 16#12;   // Connection ID for modbus Xcut #3
   "DGLASSSEARCHMACHINEINDEX_XCUT1_Q0" : DInt := 0;   // Glass search machine xcut1 quality 0
   "DGLASSSEARCHMACHINEINDEX_XCUT2_Q0" : DInt := 3;   // Glass search machine xcut2 quality 0
   "DGLASSSEARCHMACHINEINDEX_XCUT1_Q1" : DInt := 1;   // Glass search machine xcut1 quality 1
   "DGLASSSEARCHMACHINEINDEX_XCUT1_Q2" : DInt := 2;   // Glass search machine xcut1 quality 2
   "DGLASSSEARCHMACHINEINDEX_XCUT2_Q1" : DInt := 4;   // Glass search machine xcut2 quality 1
   "DGLASSSEARCHMACHINEINDEX_XCUT2_Q2" : DInt := 5;   // Glass search machine xcut2 quality 2
   "DMACHINEINDEX_GETGLASSBREAK_WANDER" : DInt := 11;   // Index get glass break data Wander Camera
   "DMAXGROSSWANDER_CMM" : DInt := 20000;   // Maximum gross wander [mm/100]
   "DMINGROSSWANDER_CMM" : DInt := -20000;   // Minimum gross wander [mm/100]
   "DMAXNETWANDER_CMM" : DInt := 20000;   // Maximum net wander [mm/100]
   "DMINNETWANDER_CMM" : DInt := -20000;   // Minimum net wander [mm/100]
   "CONNUOC_WANDER" : Conn_Ouc := 16#E;   // Connection ID for wander camera
   "IPV4_WANDER_IP1" : Byte := 192;   // IP_1 for wander camera
   "IPV4_WANDER_IP2" : Byte := 168;   // IP_2 for wander camera
   "IPV4_WANDER_IP3" : Byte := 100;   // IP_3 for wander camera
   "IPV4_WANDER_IP4" : Byte := 31;   // IP_4 for wander camera
   "UINT_WANDER_PORT" : UInt := 3000;   // Port for wander camera
   "DMAXGROSSWIDTH_CMM" : DInt := 400000;   // Maximum gross width [mm/100]
   "DMINGROSSWIDTH_CMM" : DInt := 260000;   // Minimum gross width [mm/100]
   "DMAXNETWIDTH_CMM" : DInt := 360000;   // Maximum net width [mm/100]
   "DMINNETWIDTH_CMM" : DInt := 250000;   // Minimum net width [mm/100]
   "DGLASSBREAKMACHINEINDEX_M212" : DInt := 3;   // Glass break machine M212_Man_insp
   "DGLASSBREAKGET_M209" : DInt := 8;   // Glass break get index (M209 FAN)
   "DQUALITYDESTMASK4" : LInt := 8589934592;   // Quality 4 destination mask [mask]
   "DGLASSSEARCHMACHINEINDEX_XCUT1_Q3" : DInt := 6;   // Glass search machine xcut1 quality 3
   "DGLASSSEARCHMACHINEINDEX_XCUT2_Q3" : DInt := 7;   // Glass search machine xcut2 quality 3
   "DMAXLITE_Z300" : DInt := 3;   // Maximum number of lites Z300
   "DGLASSSEARCHMACHINEINDEX_XCUT3_Q0" : DInt := 9;   // Glass search machine xcut3 quality 0
   "DGLASSSEARCHMACHINEINDEX_XCUT3_Q1" : DInt := 10;   // Glass search machine xcut3 quality 1
   "DGLASSSEARCHMACHINEINDEX_XCUT3_Q2" : DInt := 11;   // Glass search machine xcut3 quality 2
   "DGLASSSEARCHMACHINEINDEX_XCUT3_Q3" : DInt := 12;   // Glass search machine xcut3 quality 3
   "DGLASSBREAKMACHINEINDEX_M203" : DInt := 11;   // Glass break machine M203_EMXcut
   "DGLASSBREAKMACHINEINDEX_M201" : DInt := 12;   // Glass break machine M201_Snap_on_M201
   "DGLASSBREAKGET_M203" : DInt := 9;   // Glass break get index (M203 EM_XCUT)
   "DGLASSBREAKGET_M204" : DInt := 2;   // Glass break get index (M204 DropConv)
END_VAR

// folder: 01_Defects

TYPE "UDT_DefectDataExt"
TITLE = Defect data in extended mode
// Data of defect in extended mode. These defect will be sent to optimizer and reporting system.
   STRUCT
      dID : DInt;   // Defect ID [Num]
      dClass : DInt;   // Defect class value [Num]
      dSubType : DInt;   // Defect subtype [Num]
      dXPosition_cmm : DInt;   // Defect X position [mm/100]
      dYPosition_cmm : DInt;   // Defect Y position [mm/100]
      dTotalLength_um : DInt;   // Defect total length [um]
      dTotalWidth_um : DInt;   // Defect total width [um]
      dCoreLength_um : DInt;   // Defect core length [um]
      dCoreWidth_um : DInt;   // Defect core width [um]
      dDistLength_um : DInt;   // Defect distortion length [um]
      dDistWidth_um : DInt;   // Defect distortion width [um]
      dOptValue_mdptr : DInt;   // Defect optical value [mdptr]
      strDefectID : String["DSTRSIZEDEFID"];   // Defect univoque ID [string]
   END_STRUCT;
END_TYPE

TYPE "UDT_DefectData_Tracking_Ext"
TITLE = Container defect data in extended mode
// Container of defect data in extended mode. These defect will be sent to optimizer and reporting system.
   STRUCT
      dBufferHead : DInt := -1;   // Head of the buffer defect
      dBufferTail : DInt := -1;   // Tail of the buffer defect
      dBufferTailOptPLC : DInt;   // Tail plc optimizer of the buffer defect
      dBufferTailOptimizer : DInt := -1;   // Tail optimizer of the buffer defect
      dBufferTailReport : DInt := -1;   // Tail report of the buffer defect
      dDefectNextID : DInt := 1;   // Defect next ID
      xOptimizerPLCRequireAllDef : Bool;   // Optimizer plc require to resend all defects
      xOptimizerRequireAllDef : Bool := false;   // Optimizer require to resend all defects
      xBPSARequireAllDef : Bool := false;   // BPS A require to resend all defects
      xBPSBRequireAllDef : Bool;   // BPS B require to resend all defects
      rgtDefects : Array[0.."DNUMDEFEXT_IND"] of "UDT_DefectDataExt";   // Defect tank
      tDefectsForReport : Struct   // Defects structure for report
         dNumberOfDefect : DInt;   // Number of available defect
         rgtDefects : Array[0.."DNUMDEFFORREPORT_IND"] of "UDT_DefectDataExt";   // Defect tank
      END_STRUCT;
      tDefectsForOpt : Struct   // Defects structure for opt
         dNumberOfDefect : DInt;   // Number of available defect
         rgtDefects : Array[0.."DNUMDEFFOROPT_IND"] of "UDT_DefectDataExt";   // Defect tank
      END_STRUCT;
      tDefectsforOptPlc : Struct
         dNumberOfDefect : DInt;   // Number of available defect
         rgtDefects : Array[0.."DNUMDEFFOROPT_IND"] of "UDT_DefectDataExt";   // Defect tank
      END_STRUCT;
   END_STRUCT;
END_TYPE

TYPE "UDT_DefectDataRedu"
TITLE = Defect data in reducted mode
// Data of defect in reducted mode. These defect will be used from optimizer.
   STRUCT
      dClass : USInt;   // Defect class value [Num]
      dSubType : USInt;   // Defect subtype [Num]
      dXPosition_cmm : DInt;   // Defect X position [mm/100]
      dYPosition_cmm : DInt;   // Defect Y position [mm/100]
      dTotalLength_um : DInt;   // Defect total length [um]
      dTotalWidth_um : DInt;   // Defect total width [um]
   END_STRUCT;
END_TYPE

TYPE "UDT_DefectData_Tracking_Redu"
TITLE = Container defect data in reduction mode
// Container of defect data in reduction mode. These defect will be used by the internal optimizer
   STRUCT
      rgtDefClass : Array[0.."DMAXNUMCLASS_IND"] of Struct
         dBufferHead : DInt;   // Head of the buffer defect
         dBufferTail : DInt;   // Tail of the buffer defect
         tDefects : Array[0.."DMAXNUMDEFCLASS_IND"] of "UDT_DefectDataRedu";
      END_STRUCT;
   END_STRUCT;
END_TYPE

// folder: 02_Plates

TYPE "UDT_CapData"
   STRUCT
      dID : DInt;   // Cap ID [mm/100]
      dHeadPositionBTC : DInt;   // Plate head position BTC [counter]
      dTailPositionBTC : DInt;   // Plate tail position BTC [counter]
      dLength_cmm : DInt;   // Cap length [mm/100]
      dWidth_cmm : DInt;   // Cap total width [mm/100]
      dThick_cmm : DInt;   // Cap thickness [mm/100]
      dIndex : DInt;   // Cap index number in convoy [Num] (0=First cap in convoy)
      dFormat : DInt;   // Plate format [Num] (1=JS 2=Les 3=SSS)
      dNumLites : DInt;   // Number of lites in cap [Num]
      dReqGapForConv_cmm : DInt;   // Request gap beetween caps for convoy creation [mm/100]
      dMaxCapInConv : DInt;   // Maximum number of cap in convoy
      dConvTotLength_cmm : DInt;   // Total length of the convoy [mm/100]
      dMinWidth_cmm : DInt;   // Shortest width in use [mm/100]
      dMaxWidth_cmm : DInt;   // Biggest width in use [mm/100]
      dGrossWidth_cmm : DInt;   // Cap gross width [mm/100]
      dNetWidth_cmm : DInt;   // Cap net width [mm/100]
      dDEdgeOpSide_cmm : DInt;   // Double edge dimension - operator side [mm/100]
      dDEdgeOppOpSide_cmm : DInt;   // Double edge dimension - opposite operator side [mm/100]
      dTEdgeOpSide_cmm : DInt;   // Triple edge dimension - operator side [mm/100]
      dTEdgeOppOpSide_cmm : DInt;   // Triple edge dimension - opposite operator side [mm/100]
      dStartCutWander_cmm : DInt;   // Start cut wander [mm/100]
      dEndCutWander_cmm : DInt;   // End cut wander [mm/100]
      dNetWander_cmm : DInt;   // Net wander [mm/100]
      dGrossWander_cmm : DInt;   // Gross wander [mm/100]
      dColor : DInt;   // Color code [Num]
      strColorDescr : String["DSTRSIZEDESCR"];   // Color description [Text]
      dSystemMeasure : DInt;   // System of measurement (0=Metric 1=Imperial)
      tRequests : Struct   // Lavoration request on cap
         tYCutsData : Array[0.."DMAXYCUTBRIDGE_IND"] of Struct   // Requests for YCut
            xUseThisBridge : Bool;   // Use this bridge for cut
            rgdHeadsPositions : Array[0.."DMAXYHEADS_IND"] of DInt;   // Head request postions [mm/100]
            rgxHeadsRequest : Array[0.."DMAXYHEADS_IND"] of Bool;   // Head mask requests
         END_STRUCT;
         rgxXCutReqHead : Array[0.."DMAXXHEADS_IND"] of Bool;   // Request XCut Head
         rgxXCutReqTail : Array[0.."DMAXXHEADS_IND"] of Bool;   // Request XCut Tail
         rgbXCutPrioSelect : Array[0.."DMAXXHEADS_IND"] of Byte;   // Request XCut by priority manager
         xOptSelvedgeSel : Bool;   // Optimizer selvedge selection
         xOptSplitBarSel : Bool;   // Optimizer split bar selection
         xOptSepRollSel : Bool;   // Optimizer separator roll selection
         dReqTrim3OpSide : DInt;   // Request trim 3 op. side (Triple edge) with trim wheel number [x=Num]
         dReqTrim2OpSide : DInt;   // Request trim 2 op. side (Triple edge) with trim wheel number [x=Num]
         dReqTrim1OpSide : DInt;   // Request trim 1 op. side (Triple edge) with trim wheel number [x=Num]
         dReqTrim3OppOpSide : DInt;   // Request trim 3 Oppo. op. side (Triple edge) with trim wheel number [x=Num]
         dReqTrim2OppOpSide : DInt;   // Request trim 2 Oppo. op. side (Triple edge) with trim wheel number [x=Num]
         dReqTrim1OppOpSide : DInt;   // Request trim 1 Oppo. op. side (Triple edge) with trim wheel number [x=Num]
         rgdReqSplitBarSel : Array[0.."DMAXLITE_IND"] of DInt;   // Request split bar on internal cut bar number [Num]
         rgbSeparatorSelect : Array[0.."DMAXSEPROLLBANK_IND"] of Byte;   // Request separator roll mask. 1 byte each bank
         xUpdateDataBPSA : Bool;   // Request send the plate data to BPS server A
         xUpdateDataBPSB : Bool;   // Request send the plate data to BPS server B
         xWandContinue : Bool;   // Plate generated with wander in continue
         xYCutSampleTest : Bool;   // YCut sample test
         xIsCapFixed : Bool;   // Is a fixed cap
      END_STRUCT;
      tDone : Struct   // Lavoration done on cap
         tYCuts : Array[0.."DMAXYCUTBRIDGE_IND"] of Struct   // Cut done for YCut
            rgxHeadsDone : Array[0.."DMAXYHEADS_IND"] of Bool;   // Head mask done
         END_STRUCT;
         rgxXCutDoneHead : Array[0.."DMAXXHEADS_IND"] of Bool;   // Done XCut head
         rgxXCutDoneTail : Array[0.."DMAXXHEADS_IND"] of Bool;   // Done XCut tail
         xXCutDoneHead : Bool;   // XCut head cut done
         xXCutDoneTail : Bool;   // XCut tail cut done
      END_STRUCT;
      dFixedCapProductionID : DInt;   // Fixed cap production ID
      rgtLites : Array[0.."DMAXLITE_IND"] of Struct   // Lites data
         dID : DInt;   // Lite ID [Num]
         dProductionID : DInt;   // Production ID [Num]
         strProdDescr : String["DSTRSIZEDESCR"];   // Production description [Text]
         dQualityID : DInt;   // Quality ID [Num]
         strQualityDescr : String["DSTRSIZEDESCR"];   // Quality description [Text]
         dCameraRecipeID : DInt;   // Camera recipe ID [Num]
         dWidth_cmm : DInt;   // Width [mm/100]
         dBarycentre_cmm : DInt;   // Barycentre [mm/100]
         dCulletCause : DInt;   // Cullet cause
         rgxLayers : Array[0.."DMAXPROTLAYER_IND"] of Bool;   // Protection layers requested
         dMainDestination : LInt;   // Main destinations
         dAltDestination : LInt;   // Alternative destinations
         d2ndDestionation : LInt;   // Second choice destinations
         tRequests : Struct   // Request for lites
            xGeomInsp : Bool;   // Geometrical inspection request
            dMapLaserHeadOp : DInt;   // Maplaser head to print operator side [Num] (0=No print request)
            dMapLaserHeadOppOp : DInt;   // Maplaser head to print opposite operator side [Num] (0=No print request)
         END_STRUCT;
         tDone : Struct   // Done for lites
            xMapLaserHeadOp : DInt;   // Maplaser head to print operator side [Num] (0=Print not done)
            xMapLaserHeadOppOp : DInt;   // Maplaser head to print opposite operator side [Num] (0=Print not done)
         END_STRUCT;
         xSaturationPlate : Bool;   // Saturation plate
      END_STRUCT;
   END_STRUCT;
   // // rgtLites[0].rgxLayers[0] : Powder machine #1
   // // rgtLites[0].rgxLayers[1] : Powder machine #2
   // // rgtLites[0].rgxLayers[2] : Paper machine #1
END_TYPE
